(* Logix 5000 project; controller TemplateV1R0 vendor 1 type 14 code 222 rev 33.11; software revision 33.00; part 5 of 5 *)
(* UnitX_EMXXX, continued *)

ROUTINE _OM_Request_IN   (* ladder *)
// OperationMode Request
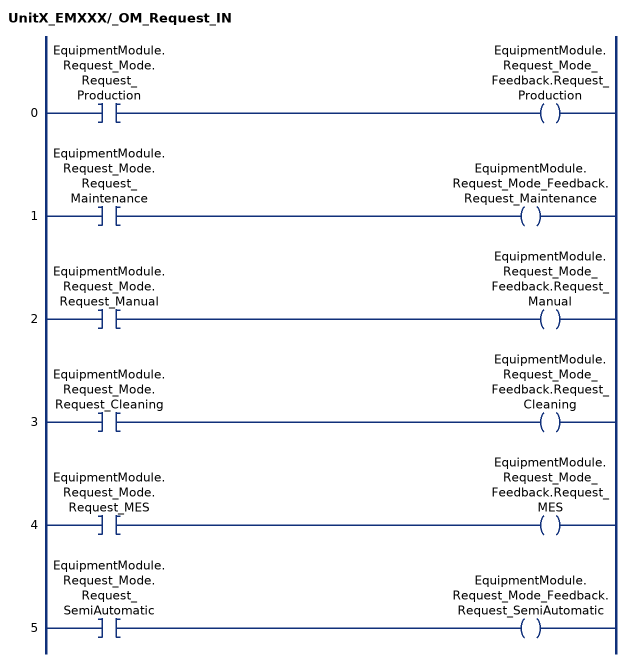
   0: XIC(EquipmentModule.Request_Mode.Request_Production)OTE(EquipmentModule.Request_Mode_Feedback.Request_Production);
   1: XIC(EquipmentModule.Request_Mode.Request_Maintenance)OTE(EquipmentModule.Request_Mode_Feedback.Request_Maintenance);
   2: XIC(EquipmentModule.Request_Mode.Request_Manual)OTE(EquipmentModule.Request_Mode_Feedback.Request_Manual);
   3: XIC(EquipmentModule.Request_Mode.Request_Cleaning)OTE(EquipmentModule.Request_Mode_Feedback.Request_Cleaning);
   4: XIC(EquipmentModule.Request_Mode.Request_MES)OTE(EquipmentModule.Request_Mode_Feedback.Request_MES);
   5: XIC(EquipmentModule.Request_Mode.Request_SemiAutomatic)OTE(EquipmentModule.Request_Mode_Feedback.Request_SemiAutomatic);
END_ROUTINE

ROUTINE Main   (* ladder *)
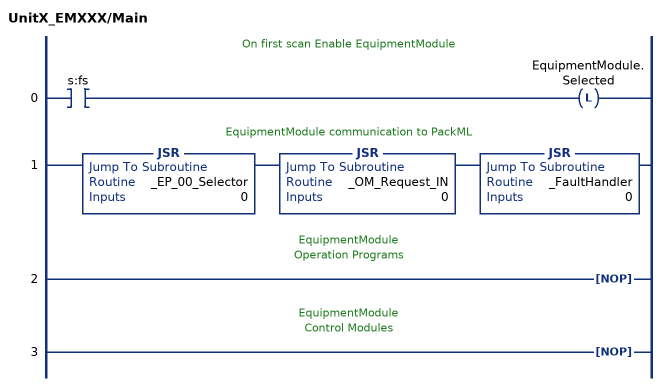
   // On first scan Enable EquipmentModule
   0: XIC(s:fs)OTL(EquipmentModule.Selected);
   // EquipmentModule communication to PackML
   1: JSR(_EP_00_Selector,0)JSR(_OM_Request_IN,0)JSR(_FaultHandler,0);
   // EquipmentModule
   // Operation Programs
   2: NOP();
   // EquipmentModule
   // Control Modules
   3: NOP();
END_ROUTINE
END_PROGRAM
